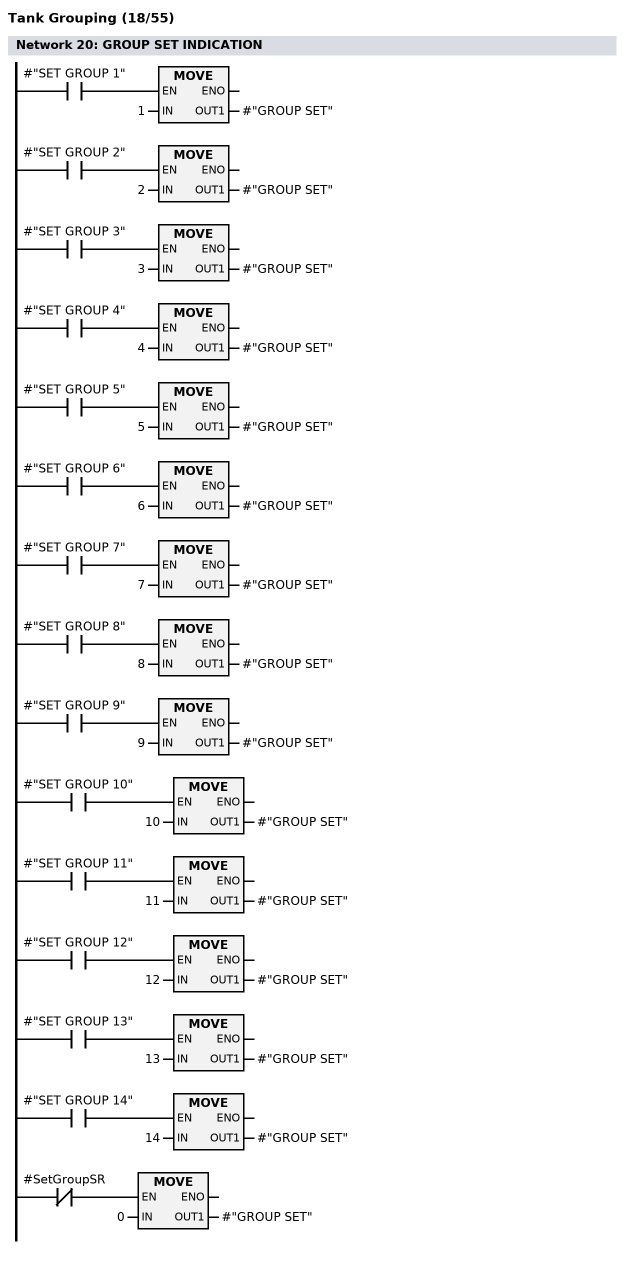
   RUNG wire#powerrail
      Contact( #"SET GROUP 1" )
      Move(in := 1, out1 => #"GROUP SET")
   END_RUNG
   RUNG wire#powerrail
      Contact( #"SET GROUP 2" )
      Move(in := 2, out1 => #"GROUP SET")
   END_RUNG
   RUNG wire#powerrail
      Contact( #"SET GROUP 3" )
      Move(in := 3, out1 => #"GROUP SET")
   END_RUNG
   RUNG wire#powerrail
      Contact( #"SET GROUP 4" )
      Move(in := 4, out1 => #"GROUP SET")
   END_RUNG
   RUNG wire#powerrail
      Contact( #"SET GROUP 5" )
      Move(in := 5, out1 => #"GROUP SET")
   END_RUNG
   RUNG wire#powerrail
      Contact( #"SET GROUP 6" )
      Move(in := 6, out1 => #"GROUP SET")
   END_RUNG
   RUNG wire#powerrail
      Contact( #"SET GROUP 7" )
      Move(in := 7, out1 => #"GROUP SET")
   END_RUNG
   RUNG wire#powerrail
      Contact( #"SET GROUP 8" )
      Move(in := 8, out1 => #"GROUP SET")
   END_RUNG
   RUNG wire#powerrail
      Contact( #"SET GROUP 9" )
      Move(in := 9, out1 => #"GROUP SET")
   END_RUNG
   RUNG wire#powerrail
      Contact( #"SET GROUP 10" )
      Move(in := 10, out1 => #"GROUP SET")
   END_RUNG
   RUNG wire#powerrail
      Contact( #"SET GROUP 11" )
      Move(in := 11, out1 => #"GROUP SET")
   END_RUNG
   RUNG wire#powerrail
      Contact( #"SET GROUP 12" )
      Move(in := 12, out1 => #"GROUP SET")
   END_RUNG
   RUNG wire#powerrail
      Contact( #"SET GROUP 13" )
      Move(in := 13, out1 => #"GROUP SET")
   END_RUNG
   RUNG wire#powerrail
      Contact( #"SET GROUP 14" )
      Move(in := 14, out1 => #"GROUP SET")
   END_RUNG
   RUNG wire#powerrail
      I_Contact( #SetGroupSR )
      Move(in := 0, out1 => #"GROUP SET")
   END_RUNG
   // the same network as SCL:
   IF #"SET GROUP 1" THEN #"GROUP SET" := 1; END_IF;
   IF #"SET GROUP 2" THEN #"GROUP SET" := 2; END_IF;
   IF #"SET GROUP 3" THEN #"GROUP SET" := 3; END_IF;
   IF #"SET GROUP 4" THEN #"GROUP SET" := 4; END_IF;
   IF #"SET GROUP 5" THEN #"GROUP SET" := 5; END_IF;
   IF #"SET GROUP 6" THEN #"GROUP SET" := 6; END_IF;
   IF #"SET GROUP 7" THEN #"GROUP SET" := 7; END_IF;
   IF #"SET GROUP 8" THEN #"GROUP SET" := 8; END_IF;
   IF #"SET GROUP 9" THEN #"GROUP SET" := 9; END_IF;
   IF #"SET GROUP 10" THEN #"GROUP SET" := 10; END_IF;
   IF #"SET GROUP 11" THEN #"GROUP SET" := 11; END_IF;
   IF #"SET GROUP 12" THEN #"GROUP SET" := 12; END_IF;
   IF #"SET GROUP 13" THEN #"GROUP SET" := 13; END_IF;
   IF #"SET GROUP 14" THEN #"GROUP SET" := 14; END_IF;
   IF NOT #SetGroupSR THEN #"GROUP SET" := 0; END_IF;
END_REGION

REGION Network 21: GROUP 1 of TANKS
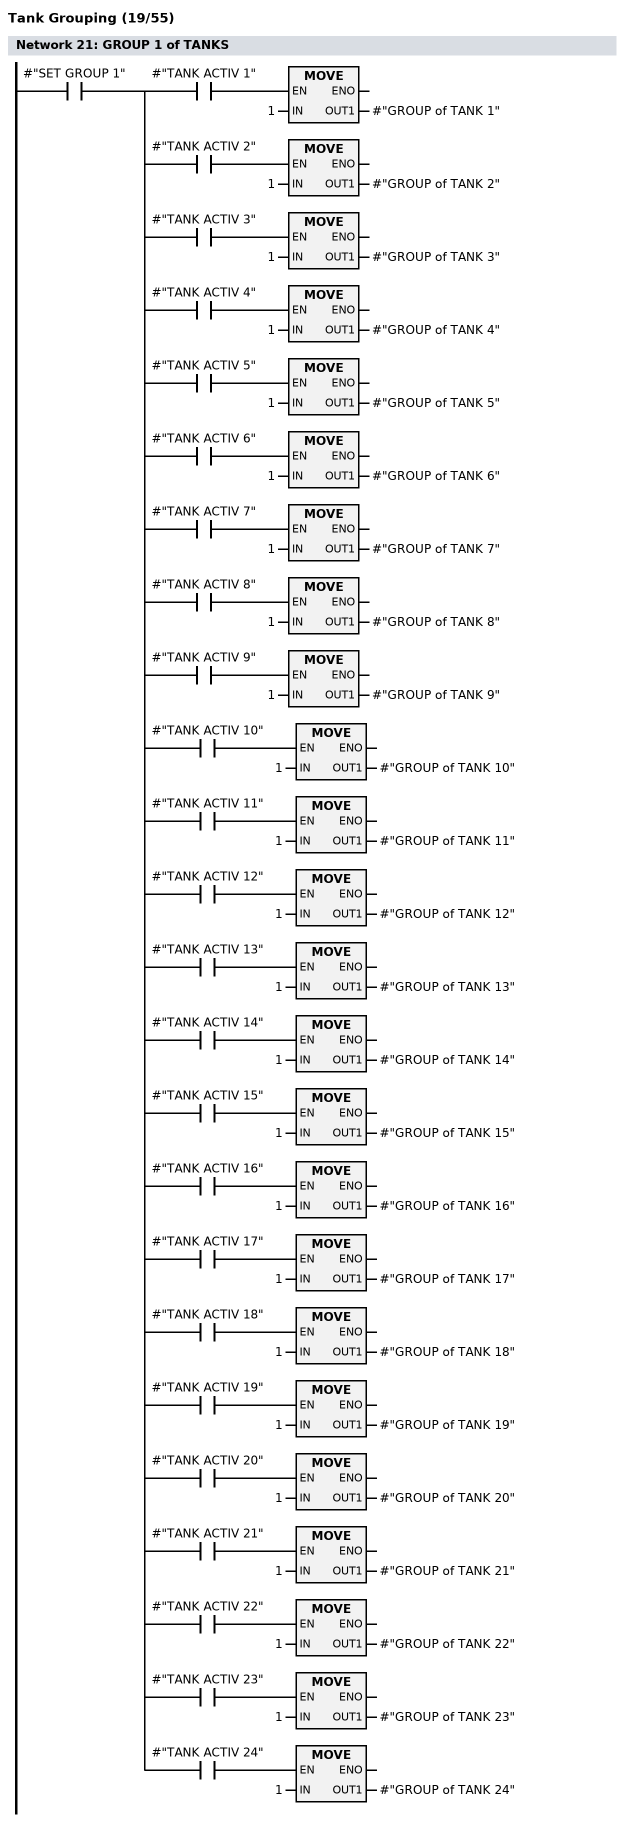
   RUNG wire#powerrail
      Contact( #"SET GROUP 1" )
      wire#w1
      Contact( #"TANK ACTIV 1" )
      Move(in := 1, out1 => #"GROUP of TANK 1")
   END_RUNG
   RUNG wire#w1
      Contact( #"TANK ACTIV 2" )
      Move(in := 1, out1 => #"GROUP of TANK 2")
   END_RUNG
   RUNG wire#w1
      Contact( #"TANK ACTIV 3" )
      Move(in := 1, out1 => #"GROUP of TANK 3")
   END_RUNG
   RUNG wire#w1
      Contact( #"TANK ACTIV 4" )
      Move(in := 1, out1 => #"GROUP of TANK 4")
   END_RUNG
   RUNG wire#w1
      Contact( #"TANK ACTIV 5" )
      Move(in := 1, out1 => #"GROUP of TANK 5")
   END_RUNG
   RUNG wire#w1
      Contact( #"TANK ACTIV 6" )
      Move(in := 1, out1 => #"GROUP of TANK 6")
   END_RUNG
   RUNG wire#w1
      Contact( #"TANK ACTIV 7" )
      Move(in := 1, out1 => #"GROUP of TANK 7")
   END_RUNG
   RUNG wire#w1
      Contact( #"TANK ACTIV 8" )
      Move(in := 1, out1 => #"GROUP of TANK 8")
   END_RUNG
   RUNG wire#w1
      Contact( #"TANK ACTIV 9" )
      Move(in := 1, out1 => #"GROUP of TANK 9")
   END_RUNG
   RUNG wire#w1
      Contact( #"TANK ACTIV 10" )
      Move(in := 1, out1 => #"GROUP of TANK 10")
   END_RUNG
   RUNG wire#w1
      Contact( #"TANK ACTIV 11" )
      Move(in := 1, out1 => #"GROUP of TANK 11")
   END_RUNG
   RUNG wire#w1
      Contact( #"TANK ACTIV 12" )
      Move(in := 1, out1 => #"GROUP of TANK 12")
   END_RUNG
   RUNG wire#w1
      Contact( #"TANK ACTIV 13" )
      Move(in := 1, out1 => #"GROUP of TANK 13")
   END_RUNG
   RUNG wire#w1
      Contact( #"TANK ACTIV 14" )
      Move(in := 1, out1 => #"GROUP of TANK 14")
   END_RUNG
   RUNG wire#w1
      Contact( #"TANK ACTIV 15" )
      Move(in := 1, out1 => #"GROUP of TANK 15")
   END_RUNG
   RUNG wire#w1
      Contact( #"TANK ACTIV 16" )
      Move(in := 1, out1 => #"GROUP of TANK 16")
   END_RUNG
   RUNG wire#w1
      Contact( #"TANK ACTIV 17" )
      Move(in := 1, out1 => #"GROUP of TANK 17")
   END_RUNG
   RUNG wire#w1
      Contact( #"TANK ACTIV 18" )
      Move(in := 1, out1 => #"GROUP of TANK 18")
   END_RUNG
   RUNG wire#w1
      Contact( #"TANK ACTIV 19" )
      Move(in := 1, out1 => #"GROUP of TANK 19")
   END_RUNG
   RUNG wire#w1
      Contact( #"TANK ACTIV 20" )
      Move(in := 1, out1 => #"GROUP of TANK 20")
   END_RUNG
   RUNG wire#w1
      Contact( #"TANK ACTIV 21" )
      Move(in := 1, out1 => #"GROUP of TANK 21")
   END_RUNG
   RUNG wire#w1
      Contact( #"TANK ACTIV 22" )
      Move(in := 1, out1 => #"GROUP of TANK 22")
   END_RUNG
   RUNG wire#w1
      Contact( #"TANK ACTIV 23" )
      Move(in := 1, out1 => #"GROUP of TANK 23")
   END_RUNG
   RUNG wire#w1
      Contact( #"TANK ACTIV 24" )
      Move(in := 1, out1 => #"GROUP of TANK 24")
   END_RUNG
   // the same network as SCL:
   IF #"SET GROUP 1" AND #"TANK ACTIV 1" THEN #"GROUP of TANK 1" := 1; END_IF;
   IF #"SET GROUP 1" AND #"TANK ACTIV 2" THEN #"GROUP of TANK 2" := 1; END_IF;
   IF #"SET GROUP 1" AND #"TANK ACTIV 3" THEN #"GROUP of TANK 3" := 1; END_IF;
   IF #"SET GROUP 1" AND #"TANK ACTIV 4" THEN #"GROUP of TANK 4" := 1; END_IF;
   IF #"SET GROUP 1" AND #"TANK ACTIV 5" THEN #"GROUP of TANK 5" := 1; END_IF;
   IF #"SET GROUP 1" AND #"TANK ACTIV 6" THEN #"GROUP of TANK 6" := 1; END_IF;
   IF #"SET GROUP 1" AND #"TANK ACTIV 7" THEN #"GROUP of TANK 7" := 1; END_IF;
   IF #"SET GROUP 1" AND #"TANK ACTIV 8" THEN #"GROUP of TANK 8" := 1; END_IF;
   IF #"SET GROUP 1" AND #"TANK ACTIV 9" THEN #"GROUP of TANK 9" := 1; END_IF;
   IF #"SET GROUP 1" AND #"TANK ACTIV 10" THEN #"GROUP of TANK 10" := 1; END_IF;
   IF #"SET GROUP 1" AND #"TANK ACTIV 11" THEN #"GROUP of TANK 11" := 1; END_IF;
   IF #"SET GROUP 1" AND #"TANK ACTIV 12" THEN #"GROUP of TANK 12" := 1; END_IF;
   IF #"SET GROUP 1" AND #"TANK ACTIV 13" THEN #"GROUP of TANK 13" := 1; END_IF;
   IF #"SET GROUP 1" AND #"TANK ACTIV 14" THEN #"GROUP of TANK 14" := 1; END_IF;
   IF #"SET GROUP 1" AND #"TANK ACTIV 15" THEN #"GROUP of TANK 15" := 1; END_IF;
   IF #"SET GROUP 1" AND #"TANK ACTIV 16" THEN #"GROUP of TANK 16" := 1; END_IF;
   IF #"SET GROUP 1" AND #"TANK ACTIV 17" THEN #"GROUP of TANK 17" := 1; END_IF;
   IF #"SET GROUP 1" AND #"TANK ACTIV 18" THEN #"GROUP of TANK 18" := 1; END_IF;
   IF #"SET GROUP 1" AND #"TANK ACTIV 19" THEN #"GROUP of TANK 19" := 1; END_IF;
   IF #"SET GROUP 1" AND #"TANK ACTIV 20" THEN #"GROUP of TANK 20" := 1; END_IF;
   IF #"SET GROUP 1" AND #"TANK ACTIV 21" THEN #"GROUP of TANK 21" := 1; END_IF;
   IF #"SET GROUP 1" AND #"TANK ACTIV 22" THEN #"GROUP of TANK 22" := 1; END_IF;
   IF #"SET GROUP 1" AND #"TANK ACTIV 23" THEN #"GROUP of TANK 23" := 1; END_IF;
   IF #"SET GROUP 1" AND #"TANK ACTIV 24" THEN #"GROUP of TANK 24" := 1; END_IF;
END_REGION

REGION Network 22: GROUP 2 of TANKS
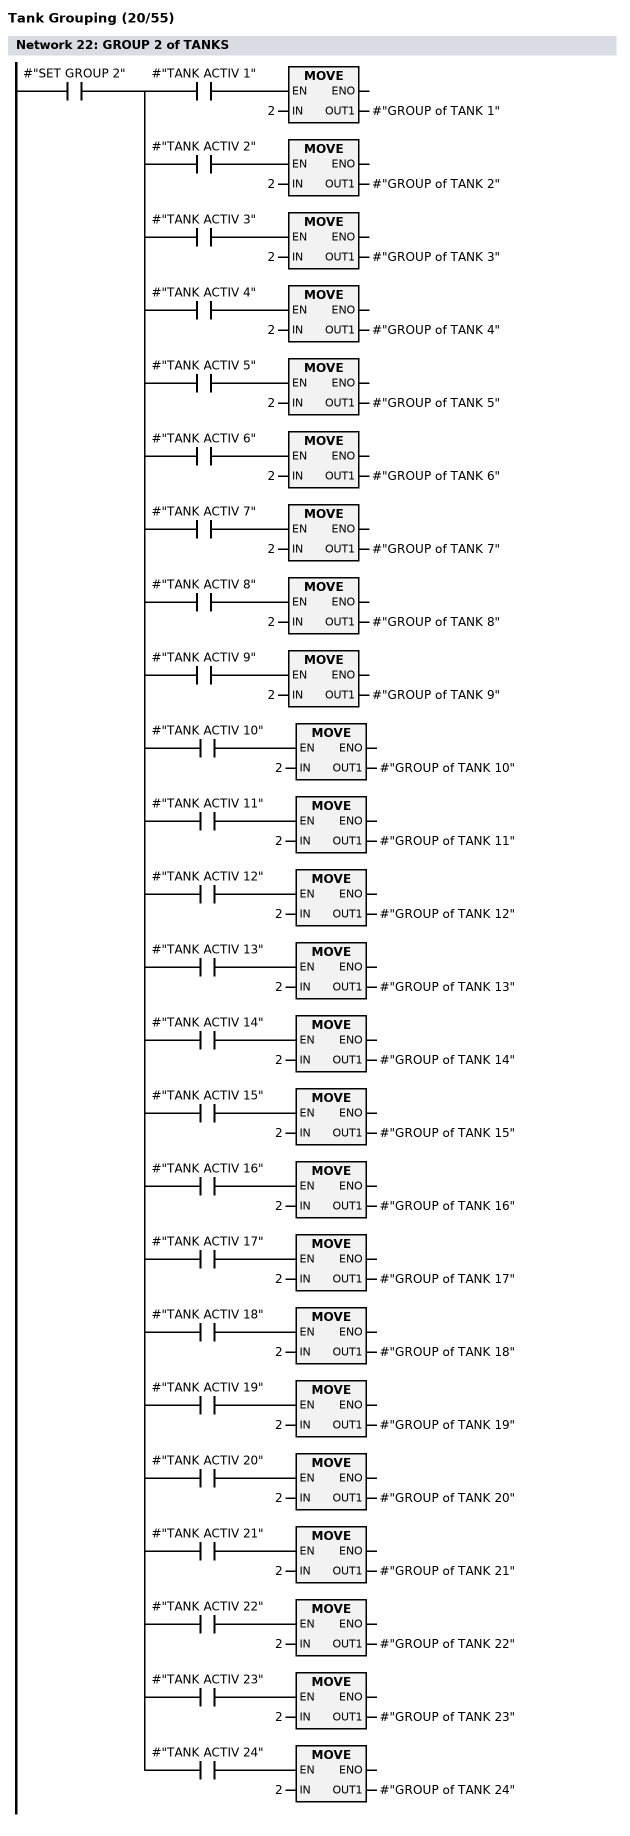
   RUNG wire#powerrail
      Contact( #"SET GROUP 2" )
      wire#w1
      Contact( #"TANK ACTIV 1" )
      Move(in := 2, out1 => #"GROUP of TANK 1")
   END_RUNG
   RUNG wire#w1
      Contact( #"TANK ACTIV 2" )
      Move(in := 2, out1 => #"GROUP of TANK 2")
   END_RUNG
   RUNG wire#w1
      Contact( #"TANK ACTIV 3" )
      Move(in := 2, out1 => #"GROUP of TANK 3")
   END_RUNG
   RUNG wire#w1
      Contact( #"TANK ACTIV 4" )
      Move(in := 2, out1 => #"GROUP of TANK 4")
   END_RUNG
   RUNG wire#w1
      Contact( #"TANK ACTIV 5" )
      Move(in := 2, out1 => #"GROUP of TANK 5")
   END_RUNG
   RUNG wire#w1
      Contact( #"TANK ACTIV 6" )
      Move(in := 2, out1 => #"GROUP of TANK 6")
   END_RUNG
   RUNG wire#w1
      Contact( #"TANK ACTIV 7" )
      Move(in := 2, out1 => #"GROUP of TANK 7")
   END_RUNG
   RUNG wire#w1
      Contact( #"TANK ACTIV 8" )
      Move(in := 2, out1 => #"GROUP of TANK 8")
   END_RUNG
   RUNG wire#w1
      Contact( #"TANK ACTIV 9" )
      Move(in := 2, out1 => #"GROUP of TANK 9")
   END_RUNG
   RUNG wire#w1
      Contact( #"TANK ACTIV 10" )
      Move(in := 2, out1 => #"GROUP of TANK 10")
   END_RUNG
   RUNG wire#w1
      Contact( #"TANK ACTIV 11" )
      Move(in := 2, out1 => #"GROUP of TANK 11")
   END_RUNG
   RUNG wire#w1
      Contact( #"TANK ACTIV 12" )
      Move(in := 2, out1 => #"GROUP of TANK 12")
   END_RUNG
   RUNG wire#w1
      Contact( #"TANK ACTIV 13" )
      Move(in := 2, out1 => #"GROUP of TANK 13")
   END_RUNG
   RUNG wire#w1
      Contact( #"TANK ACTIV 14" )
      Move(in := 2, out1 => #"GROUP of TANK 14")
   END_RUNG
   RUNG wire#w1
      Contact( #"TANK ACTIV 15" )
      Move(in := 2, out1 => #"GROUP of TANK 15")
   END_RUNG
   RUNG wire#w1
      Contact( #"TANK ACTIV 16" )
      Move(in := 2, out1 => #"GROUP of TANK 16")
   END_RUNG
   RUNG wire#w1
      Contact( #"TANK ACTIV 17" )
      Move(in := 2, out1 => #"GROUP of TANK 17")
   END_RUNG
   RUNG wire#w1
      Contact( #"TANK ACTIV 18" )
      Move(in := 2, out1 => #"GROUP of TANK 18")
   END_RUNG
   RUNG wire#w1
      Contact( #"TANK ACTIV 19" )
      Move(in := 2, out1 => #"GROUP of TANK 19")
   END_RUNG
   RUNG wire#w1
      Contact( #"TANK ACTIV 20" )
      Move(in := 2, out1 => #"GROUP of TANK 20")
   END_RUNG
   RUNG wire#w1
      Contact( #"TANK ACTIV 21" )
      Move(in := 2, out1 => #"GROUP of TANK 21")
   END_RUNG
   RUNG wire#w1
      Contact( #"TANK ACTIV 22" )
      Move(in := 2, out1 => #"GROUP of TANK 22")
   END_RUNG
   RUNG wire#w1
      Contact( #"TANK ACTIV 23" )
      Move(in := 2, out1 => #"GROUP of TANK 23")
   END_RUNG
   RUNG wire#w1
      Contact( #"TANK ACTIV 24" )
      Move(in := 2, out1 => #"GROUP of TANK 24")
   END_RUNG
   // the same network as SCL:
   IF #"SET GROUP 2" AND #"TANK ACTIV 1" THEN #"GROUP of TANK 1" := 2; END_IF;
   IF #"SET GROUP 2" AND #"TANK ACTIV 2" THEN #"GROUP of TANK 2" := 2; END_IF;
   IF #"SET GROUP 2" AND #"TANK ACTIV 3" THEN #"GROUP of TANK 3" := 2; END_IF;
   IF #"SET GROUP 2" AND #"TANK ACTIV 4" THEN #"GROUP of TANK 4" := 2; END_IF;
   IF #"SET GROUP 2" AND #"TANK ACTIV 5" THEN #"GROUP of TANK 5" := 2; END_IF;
   IF #"SET GROUP 2" AND #"TANK ACTIV 6" THEN #"GROUP of TANK 6" := 2; END_IF;
   IF #"SET GROUP 2" AND #"TANK ACTIV 7" THEN #"GROUP of TANK 7" := 2; END_IF;
   IF #"SET GROUP 2" AND #"TANK ACTIV 8" THEN #"GROUP of TANK 8" := 2; END_IF;
   IF #"SET GROUP 2" AND #"TANK ACTIV 9" THEN #"GROUP of TANK 9" := 2; END_IF;
   IF #"SET GROUP 2" AND #"TANK ACTIV 10" THEN #"GROUP of TANK 10" := 2; END_IF;
   IF #"SET GROUP 2" AND #"TANK ACTIV 11" THEN #"GROUP of TANK 11" := 2; END_IF;
   IF #"SET GROUP 2" AND #"TANK ACTIV 12" THEN #"GROUP of TANK 12" := 2; END_IF;
   IF #"SET GROUP 2" AND #"TANK ACTIV 13" THEN #"GROUP of TANK 13" := 2; END_IF;
   IF #"SET GROUP 2" AND #"TANK ACTIV 14" THEN #"GROUP of TANK 14" := 2; END_IF;
   IF #"SET GROUP 2" AND #"TANK ACTIV 15" THEN #"GROUP of TANK 15" := 2; END_IF;
   IF #"SET GROUP 2" AND #"TANK ACTIV 16" THEN #"GROUP of TANK 16" := 2; END_IF;
   IF #"SET GROUP 2" AND #"TANK ACTIV 17" THEN #"GROUP of TANK 17" := 2; END_IF;
   IF #"SET GROUP 2" AND #"TANK ACTIV 18" THEN #"GROUP of TANK 18" := 2; END_IF;
   IF #"SET GROUP 2" AND #"TANK ACTIV 19" THEN #"GROUP of TANK 19" := 2; END_IF;
   IF #"SET GROUP 2" AND #"TANK ACTIV 20" THEN #"GROUP of TANK 20" := 2; END_IF;
   IF #"SET GROUP 2" AND #"TANK ACTIV 21" THEN #"GROUP of TANK 21" := 2; END_IF;
   IF #"SET GROUP 2" AND #"TANK ACTIV 22" THEN #"GROUP of TANK 22" := 2; END_IF;
   IF #"SET GROUP 2" AND #"TANK ACTIV 23" THEN #"GROUP of TANK 23" := 2; END_IF;
   IF #"SET GROUP 2" AND #"TANK ACTIV 24" THEN #"GROUP of TANK 24" := 2; END_IF;
END_REGION

REGION Network 23: GROUP 3 of TANKS
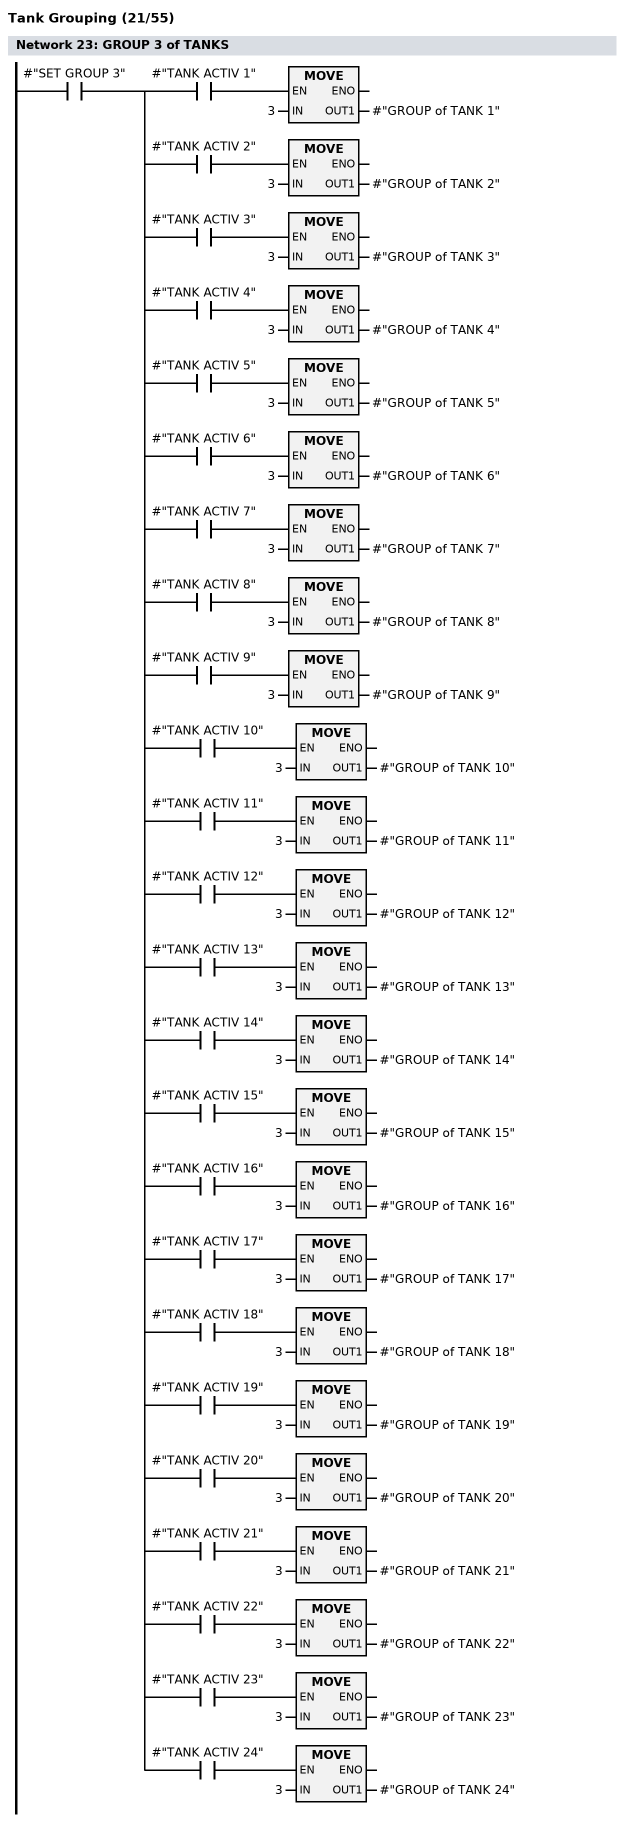
   RUNG wire#powerrail
      Contact( #"SET GROUP 3" )
      wire#w1
      Contact( #"TANK ACTIV 1" )
      Move(in := 3, out1 => #"GROUP of TANK 1")
   END_RUNG
   RUNG wire#w1
      Contact( #"TANK ACTIV 2" )
      Move(in := 3, out1 => #"GROUP of TANK 2")
   END_RUNG
   RUNG wire#w1
      Contact( #"TANK ACTIV 3" )
      Move(in := 3, out1 => #"GROUP of TANK 3")
   END_RUNG
   RUNG wire#w1
      Contact( #"TANK ACTIV 4" )
      Move(in := 3, out1 => #"GROUP of TANK 4")
   END_RUNG
   RUNG wire#w1
      Contact( #"TANK ACTIV 5" )
      Move(in := 3, out1 => #"GROUP of TANK 5")
   END_RUNG
   RUNG wire#w1
      Contact( #"TANK ACTIV 6" )
      Move(in := 3, out1 => #"GROUP of TANK 6")
   END_RUNG
   RUNG wire#w1
      Contact( #"TANK ACTIV 7" )
      Move(in := 3, out1 => #"GROUP of TANK 7")
   END_RUNG
   RUNG wire#w1
      Contact( #"TANK ACTIV 8" )
      Move(in := 3, out1 => #"GROUP of TANK 8")
   END_RUNG
   RUNG wire#w1
      Contact( #"TANK ACTIV 9" )
      Move(in := 3, out1 => #"GROUP of TANK 9")
   END_RUNG
   RUNG wire#w1
      Contact( #"TANK ACTIV 10" )
      Move(in := 3, out1 => #"GROUP of TANK 10")
   END_RUNG
   RUNG wire#w1
      Contact( #"TANK ACTIV 11" )
      Move(in := 3, out1 => #"GROUP of TANK 11")
   END_RUNG
   RUNG wire#w1
      Contact( #"TANK ACTIV 12" )
      Move(in := 3, out1 => #"GROUP of TANK 12")
   END_RUNG
   RUNG wire#w1
      Contact( #"TANK ACTIV 13" )
      Move(in := 3, out1 => #"GROUP of TANK 13")
   END_RUNG
   RUNG wire#w1
      Contact( #"TANK ACTIV 14" )
      Move(in := 3, out1 => #"GROUP of TANK 14")
   END_RUNG
   RUNG wire#w1
      Contact( #"TANK ACTIV 15" )
      Move(in := 3, out1 => #"GROUP of TANK 15")
   END_RUNG
   RUNG wire#w1
      Contact( #"TANK ACTIV 16" )
      Move(in := 3, out1 => #"GROUP of TANK 16")
   END_RUNG
   RUNG wire#w1
      Contact( #"TANK ACTIV 17" )
      Move(in := 3, out1 => #"GROUP of TANK 17")
   END_RUNG
   RUNG wire#w1
      Contact( #"TANK ACTIV 18" )
      Move(in := 3, out1 => #"GROUP of TANK 18")
   END_RUNG
   RUNG wire#w1
      Contact( #"TANK ACTIV 19" )
      Move(in := 3, out1 => #"GROUP of TANK 19")
   END_RUNG
   RUNG wire#w1
      Contact( #"TANK ACTIV 20" )
      Move(in := 3, out1 => #"GROUP of TANK 20")
   END_RUNG
   RUNG wire#w1
      Contact( #"TANK ACTIV 21" )
      Move(in := 3, out1 => #"GROUP of TANK 21")
   END_RUNG
   RUNG wire#w1
      Contact( #"TANK ACTIV 22" )
      Move(in := 3, out1 => #"GROUP of TANK 22")
   END_RUNG
   RUNG wire#w1
      Contact( #"TANK ACTIV 23" )
      Move(in := 3, out1 => #"GROUP of TANK 23")